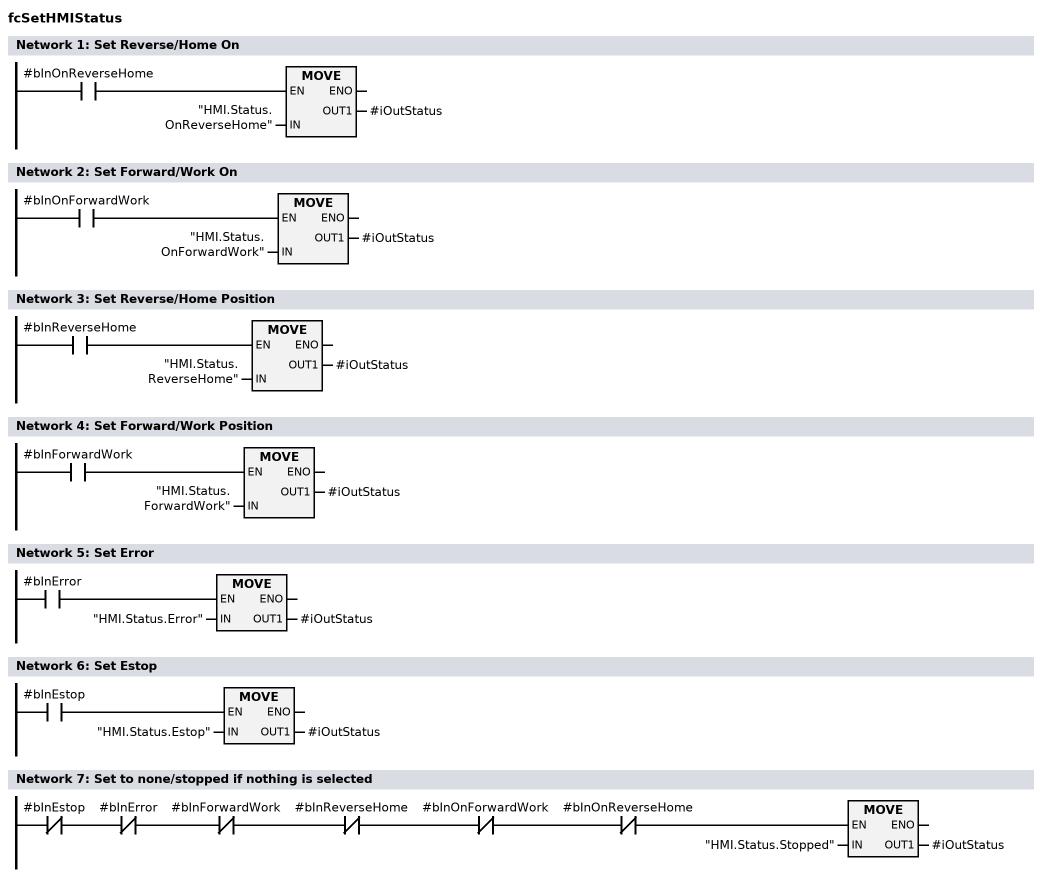
   RUNG wire#powerrail
      Contact( #bInOnReverseHome )
      Move(in := "HMI.Status.OnReverseHome", out1 => #iOutStatus)
   END_RUNG
   // the same network as SCL:
   IF #bInOnReverseHome THEN #iOutStatus := "HMI.Status.OnReverseHome"; END_IF;
END_REGION

REGION Network 2: Set Forward/Work On
   RUNG wire#powerrail
      Contact( #bInOnForwardWork )
      Move(in := "HMI.Status.OnForwardWork", out1 => #iOutStatus)
   END_RUNG
   // the same network as SCL:
   IF #bInOnForwardWork THEN #iOutStatus := "HMI.Status.OnForwardWork"; END_IF;
END_REGION

REGION Network 3: Set Reverse/Home Position
   RUNG wire#powerrail
      Contact( #bInReverseHome )
      Move(in := "HMI.Status.ReverseHome", out1 => #iOutStatus)
   END_RUNG
   // the same network as SCL:
   IF #bInReverseHome THEN #iOutStatus := "HMI.Status.ReverseHome"; END_IF;
END_REGION

REGION Network 4: Set Forward/Work Position
   RUNG wire#powerrail
      Contact( #bInForwardWork )
      Move(in := "HMI.Status.ForwardWork", out1 => #iOutStatus)
   END_RUNG
   // the same network as SCL:
   IF #bInForwardWork THEN #iOutStatus := "HMI.Status.ForwardWork"; END_IF;
END_REGION

REGION Network 5: Set Error
   RUNG wire#powerrail
      Contact( #bInError )
      Move(in := "HMI.Status.Error", out1 => #iOutStatus)
   END_RUNG
   // the same network as SCL:
   IF #bInError THEN #iOutStatus := "HMI.Status.Error"; END_IF;
END_REGION

REGION Network 6: Set Estop
   RUNG wire#powerrail
      Contact( #bInEstop )
      Move(in := "HMI.Status.Estop", out1 => #iOutStatus)
   END_RUNG
   // the same network as SCL:
   IF #bInEstop THEN #iOutStatus := "HMI.Status.Estop"; END_IF;
END_REGION

REGION Network 7: Set to none/stopped if nothing is selected
   RUNG wire#powerrail
      I_Contact( #bInEstop )
      I_Contact( #bInError )
      I_Contact( #bInForwardWork )
      I_Contact( #bInReverseHome )
      I_Contact( #bInOnForwardWork )
      I_Contact( #bInOnReverseHome )
      Move(in := "HMI.Status.Stopped", out1 => #iOutStatus)
   END_RUNG
   // the same network as SCL:
   IF NOT #bInEstop AND NOT #bInError AND NOT #bInForwardWork AND NOT #bInReverseHome AND NOT #bInOnForwardWork AND NOT #bInOnReverseHome THEN
       #iOutStatus := "HMI.Status.Stopped";
   END_IF;
END_REGION
END_FUNCTION

FUNCTION "fcSetHMIStatusGeneric" : Void   // FC1121, LAD
TITLE = Sets HMI Status
{ S7_Optimized_Access := 'FALSE' }
VERSION : 0.1
// Wrapper function for setting the HMI status of a device. 
// 
// It will display in order of priority, based on input, where Status1 > Status 2 > Status 3 > Status 4 > Status 5 > Status 6.
BEGIN

REGION Network 1: Set Status 6
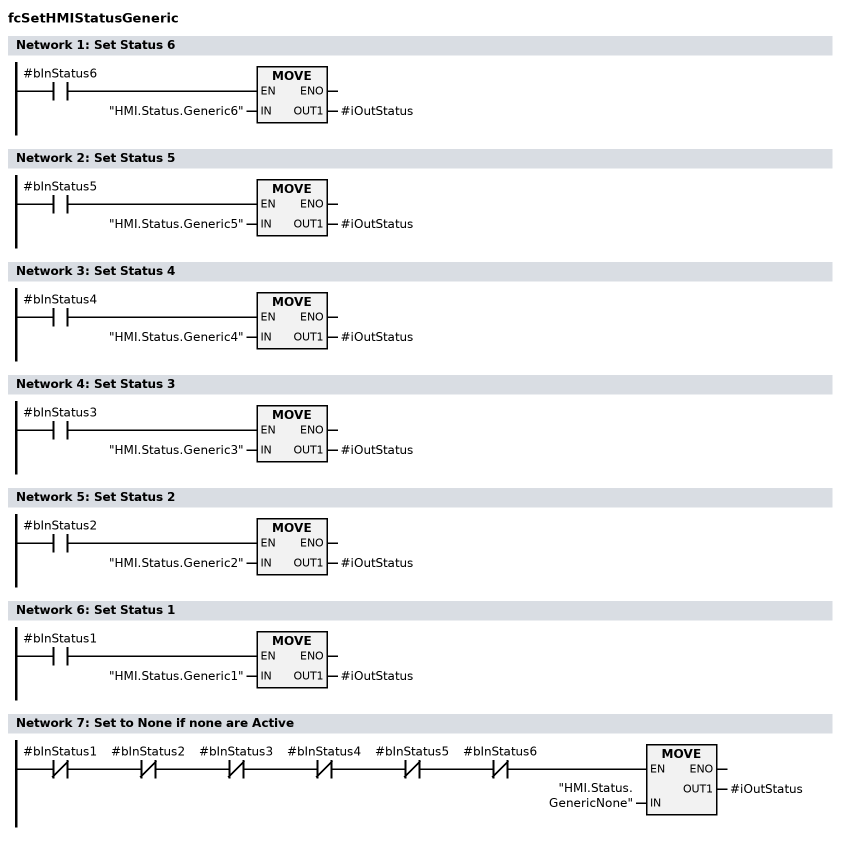
   RUNG wire#powerrail
      Contact( #bInStatus6 )
      { S7_GenerateENO := "TRUE" } Move(in := "HMI.Status.Generic6", out1 => #iOutStatus)
   END_RUNG
   // the same network as SCL:
   IF #bInStatus6 THEN #iOutStatus := "HMI.Status.Generic6"; END_IF;
END_REGION

REGION Network 2: Set Status 5
   RUNG wire#powerrail
      Contact( #bInStatus5 )
      { S7_GenerateENO := "TRUE" } Move(in := "HMI.Status.Generic5", out1 => #iOutStatus)
   END_RUNG
   // the same network as SCL:
   IF #bInStatus5 THEN #iOutStatus := "HMI.Status.Generic5"; END_IF;
END_REGION

REGION Network 3: Set Status 4
   RUNG wire#powerrail
      Contact( #bInStatus4 )
      { S7_GenerateENO := "TRUE" } Move(in := "HMI.Status.Generic4", out1 => #iOutStatus)
   END_RUNG
   // the same network as SCL:
   IF #bInStatus4 THEN #iOutStatus := "HMI.Status.Generic4"; END_IF;
END_REGION

REGION Network 4: Set Status 3
   RUNG wire#powerrail
      Contact( #bInStatus3 )
      { S7_GenerateENO := "TRUE" } Move(in := "HMI.Status.Generic3", out1 => #iOutStatus)
   END_RUNG
   // the same network as SCL:
   IF #bInStatus3 THEN #iOutStatus := "HMI.Status.Generic3"; END_IF;
END_REGION

REGION Network 5: Set Status 2
   RUNG wire#powerrail
      Contact( #bInStatus2 )
      { S7_GenerateENO := "TRUE" } Move(in := "HMI.Status.Generic2", out1 => #iOutStatus)
   END_RUNG
   // the same network as SCL:
   IF #bInStatus2 THEN #iOutStatus := "HMI.Status.Generic2"; END_IF;
END_REGION

REGION Network 6: Set Status 1
   RUNG wire#powerrail
      Contact( #bInStatus1 )
      { S7_GenerateENO := "TRUE" } Move(in := "HMI.Status.Generic1", out1 => #iOutStatus)
   END_RUNG
   // the same network as SCL:
   IF #bInStatus1 THEN #iOutStatus := "HMI.Status.Generic1"; END_IF;
END_REGION

REGION Network 7: Set to None if none are Active
   RUNG wire#powerrail
      I_Contact( #bInStatus1 )
      I_Contact( #bInStatus2 )
      I_Contact( #bInStatus3 )
      I_Contact( #bInStatus4 )
      I_Contact( #bInStatus5 )
      I_Contact( #bInStatus6 )
      { S7_GenerateENO := "TRUE" } Move(in := "HMI.Status.GenericNone", out1 => #iOutStatus)
   END_RUNG
   // the same network as SCL:
   IF NOT #bInStatus1 AND NOT #bInStatus2 AND NOT #bInStatus3 AND NOT #bInStatus4 AND NOT #bInStatus5 AND NOT #bInStatus6 THEN
       #iOutStatus := "HMI.Status.GenericNone";
   END_IF;
END_REGION
END_FUNCTION

// folder: Library Blocks/Resources/IO

FUNCTION "fcReadInput" : Void   // FC301, LAD
TITLE = Read/Scale input word
{ S7_Optimized_Access := 'FALSE' }
AUTHOR : DMC
FAMILY : IO
VERSION : 0.1
   VAR_TEMP   // added for the SCL form of the ladder/FBD networks
      _w1 : Bool;
      _w2 : Bool;
   END_VAR
BEGIN

REGION Network 1: Swap input value bytes if needed
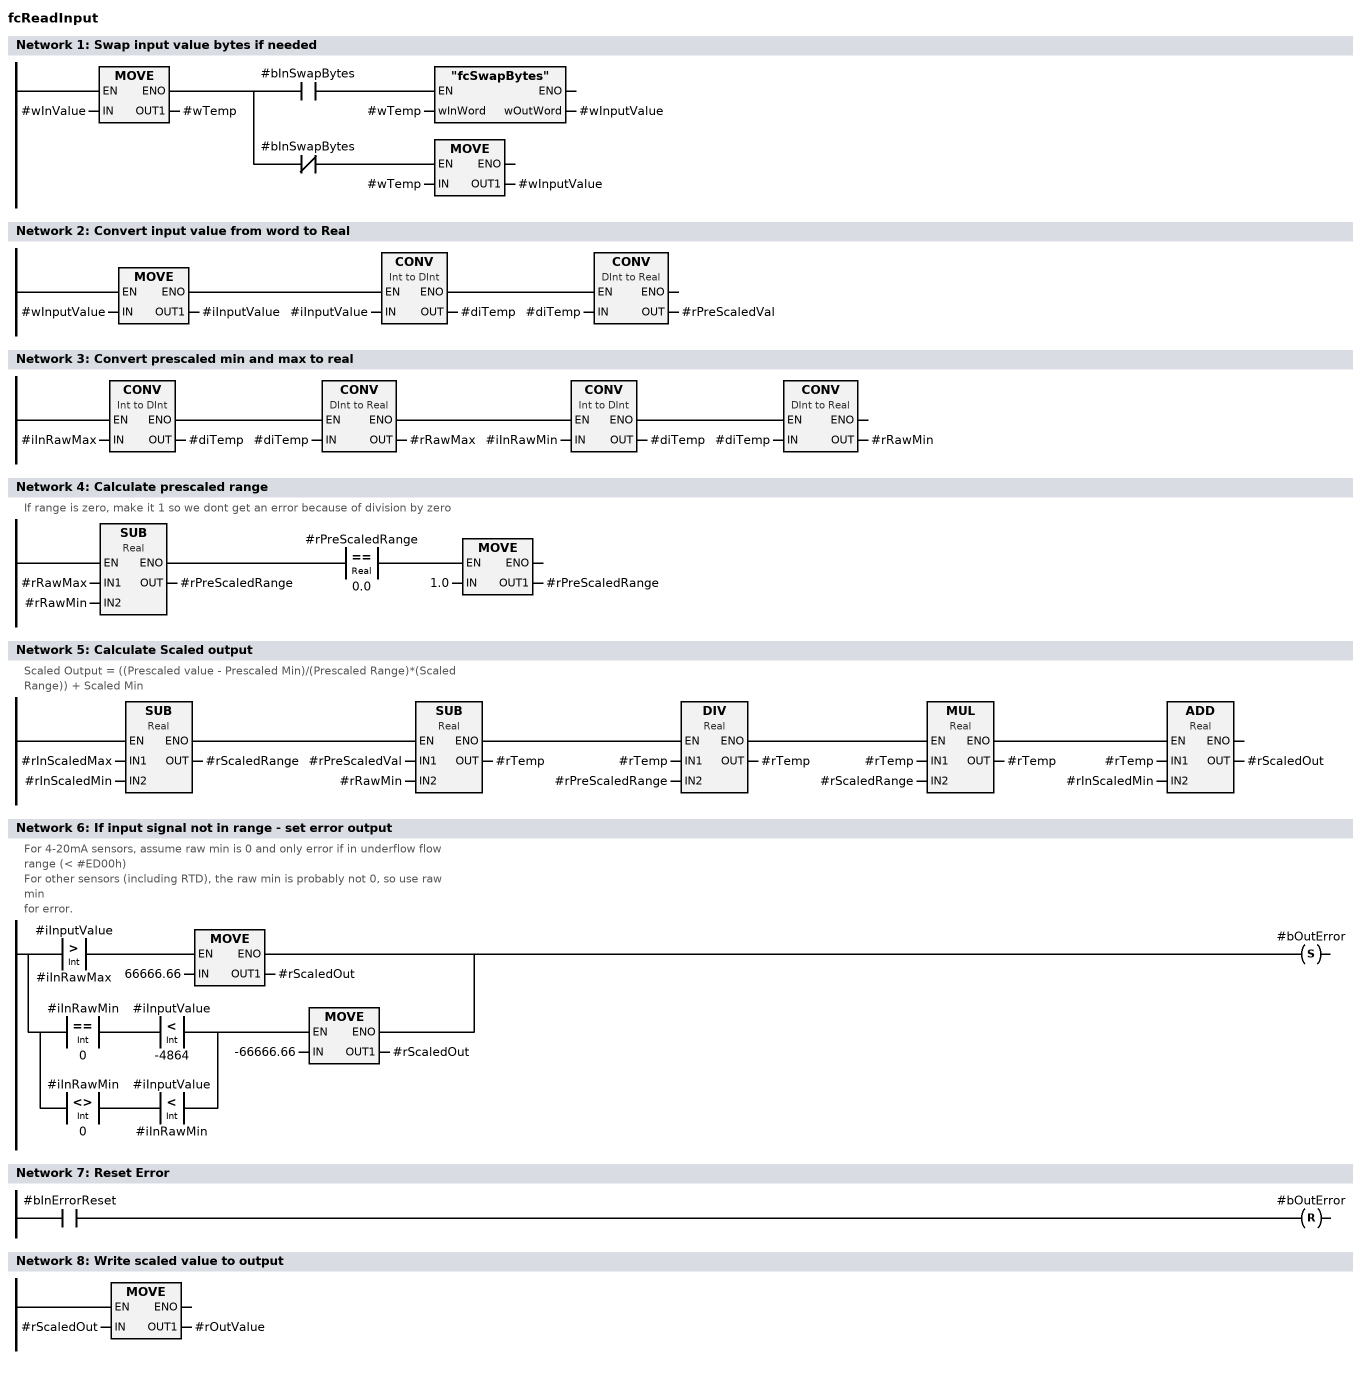
   RUNG wire#powerrail
      { S7_GenerateENO := "TRUE" } Move(in := #wInValue, out1 => #wTemp)
      wire#w1
      Contact( #bInSwapBytes )
      "fcSwapBytes"(wInWord := #wTemp, wOutWord => #wInputValue)
   END_RUNG
   RUNG wire#w1
      I_Contact( #bInSwapBytes )
      { S7_GenerateENO := "TRUE" } Move(in := #wTemp, out1 => #wInputValue)
   END_RUNG
   // the same network as SCL:
   // ENO of a box is taken as its EN; it also drops when the box reports an error
   #wTemp := #wInValue;
   IF #bInSwapBytes THEN "fcSwapBytes"(wInWord := #wTemp, wOutWord => #wInputValue); END_IF;
   IF NOT #bInSwapBytes THEN #wInputValue := #wTemp; END_IF;
END_REGION

REGION Network 2: Convert input value from word to Real
   RUNG wire#powerrail
      { S7_GenerateENO := "TRUE" } Move(in := #wInputValue, out1 => #iInputValue)
      { S7_Templates := "[SrcType := Int, DestType := DInt]"; S7_GenerateENO := "TRUE" } Convert(in := #iInputValue, out => #diTemp)
      { S7_Templates := "[SrcType := DInt, DestType := Real]"; S7_GenerateENO := "TRUE" } Convert(in := #diTemp, out => #rPreScaledVal)
   END_RUNG
   // the same network as SCL:
   // ENO of a box is taken as its EN; it also drops when the box reports an error
   #iInputValue := #wInputValue;
   #diTemp := INT_TO_DINT(#iInputValue);
   #rPreScaledVal := DINT_TO_REAL(#diTemp);
END_REGION

REGION Network 3: Convert prescaled min and max to real
   RUNG wire#powerrail
      { S7_Templates := "[SrcType := Int, DestType := DInt]"; S7_GenerateENO := "TRUE" } Convert(in := #iInRawMax, out => #diTemp)
      { S7_Templates := "[SrcType := DInt, DestType := Real]"; S7_GenerateENO := "TRUE" } Convert(in := #diTemp, out => #rRawMax)
      { S7_Templates := "[SrcType := Int, DestType := DInt]"; S7_GenerateENO := "TRUE" } Convert(in := #iInRawMin, out => #diTemp)
      { S7_Templates := "[SrcType := DInt, DestType := Real]"; S7_GenerateENO := "TRUE" } Convert(in := #diTemp, out => #rRawMin)
   END_RUNG
   // the same network as SCL:
   // ENO of a box is taken as its EN; it also drops when the box reports an error
   #diTemp := INT_TO_DINT(#iInRawMax);
   #rRawMax := DINT_TO_REAL(#diTemp);
   #diTemp := INT_TO_DINT(#iInRawMin);
   #rRawMin := DINT_TO_REAL(#diTemp);
END_REGION

REGION Network 4: Calculate prescaled range
   // If range is zero, make it 1 so we dont get an error because of division by zero
   RUNG wire#powerrail
      { S7_Templates := "SrcType := Real"; S7_GenerateENO := "TRUE" } Sub(in1 := #rRawMax, in2 := #rRawMin, out => #rPreScaledRange)
      { S7_Templates := "SrcType := Real" } EQ_Contact(in1 := #rPreScaledRange, in2 := 0.0)
      { S7_GenerateENO := "TRUE" } Move(in := 1.0, out1 => #rPreScaledRange)
   END_RUNG
   // the same network as SCL:
   // ENO of a box is taken as its EN; it also drops when the box reports an error
   #rPreScaledRange := #rRawMax - #rRawMin;
   IF #rPreScaledRange = 0.0 THEN #rPreScaledRange := 1.0; END_IF;
END_REGION

REGION Network 5: Calculate Scaled output
   // Scaled Output = ((Prescaled value - Prescaled Min)/(Prescaled Range)*(Scaled 
   // Range)) + Scaled Min
   RUNG wire#powerrail
      { S7_Templates := "SrcType := Real"; S7_GenerateENO := "TRUE" } Sub(in1 := #rInScaledMax, in2 := #rInScaledMin, out => #rScaledRange)
      { S7_Templates := "SrcType := Real"; S7_GenerateENO := "TRUE" } Sub(in1 := #rPreScaledVal, in2 := #rRawMin, out => #rTemp)
      { S7_Templates := "SrcType := Real"; S7_GenerateENO := "TRUE" } Div(in1 := #rTemp, in2 := #rPreScaledRange, out => #rTemp)
      { S7_Templates := "SrcType := Real"; S7_GenerateENO := "TRUE" } Mul(in1 := #rTemp, in2 := #rScaledRange, out => #rTemp)
      { S7_Templates := "SrcType := Real"; S7_GenerateENO := "TRUE" } Add(in1 := #rTemp, in2 := #rInScaledMin, out => #rScaledOut)
   END_RUNG
   // the same network as SCL:
   // ENO of a box is taken as its EN; it also drops when the box reports an error
   #rScaledRange := #rInScaledMax - #rInScaledMin;
   #rTemp := #rPreScaledVal - #rRawMin;
   #rTemp := #rTemp / #rPreScaledRange;
   #rTemp := #rTemp * #rScaledRange;
   #rScaledOut := #rTemp + #rInScaledMin;
END_REGION

REGION Network 6: If input signal not in range - set error output
   // For 4-20mA sensors, assume raw min is 0 and only error if in underflow flow 
   // range (< #ED00h)
   // 
   // For other sensors (including RTD), the raw min is probably not 0, so use raw 
   // min 
   // for error.
   RUNG wire#powerrail
      { S7_Templates := "SrcType := Int" } GT_Contact(in1 := #iInputValue, in2 := #iInRawMax)
      { S7_GenerateENO := "TRUE" } Move(in := 66666.66, out1 => #rScaledOut)
      wire#w1
      S_Coil( #bOutError )
   END_RUNG
   RUNG wire#powerrail
      { S7_Templates := "SrcType := Int" } EQ_Contact(in1 := #iInRawMin, in2 := 0)
      { S7_Templates := "SrcType := Int" } LT_Contact(in1 := #iInputValue, in2 := -4864)
      wire#w2
      { S7_GenerateENO := "TRUE" } Move(in := -66666.66, out1 => #rScaledOut)
   END_RUNG wire#w1
   RUNG wire#powerrail
      { S7_Templates := "SrcType := Int" } NE_Contact(in1 := #iInRawMin, in2 := 0)
      { S7_Templates := "SrcType := Int" } LT_Contact(in1 := #iInputValue, in2 := #iInRawMin)
   END_RUNG wire#w2
   // the same network as SCL:
   // ENO of a box is taken as its EN; it also drops when the box reports an error
   #_w1 := #iInputValue > #iInRawMax;
   IF #_w1 THEN #rScaledOut := 66666.66; END_IF;
   #_w2 := ((#iInRawMin = 0) AND (#iInputValue < (-4864))) OR ((#iInRawMin <> 0) AND (#iInputValue < #iInRawMin));
   IF #_w2 THEN #rScaledOut := -66666.66; END_IF;
   IF #_w1 OR #_w2 THEN #bOutError := TRUE; END_IF;
END_REGION

REGION Network 7: Reset Error
   RUNG wire#powerrail
      Contact( #bInErrorReset )
      R_Coil( #bOutError )
   END_RUNG
   // the same network as SCL:
   IF #bInErrorReset THEN #bOutError := FALSE; END_IF;
END_REGION

REGION Network 8: Write scaled value to output
   RUNG wire#powerrail
      { S7_GenerateENO := "TRUE" } Move(in := #rScaledOut, out1 => #rOutValue)
   END_RUNG
   // the same network as SCL:
   #rOutValue := #rScaledOut;
END_REGION
END_FUNCTION

FUNCTION "fcWriteOutput" : Void   // FC302, LAD
TITLE = Writes a scaled output
{ S7_Optimized_Access := 'FALSE' }
AUTHOR : DMC
FAMILY : IO
VERSION : 0.1
BEGIN

REGION Network 1: Convert raw min and max to real
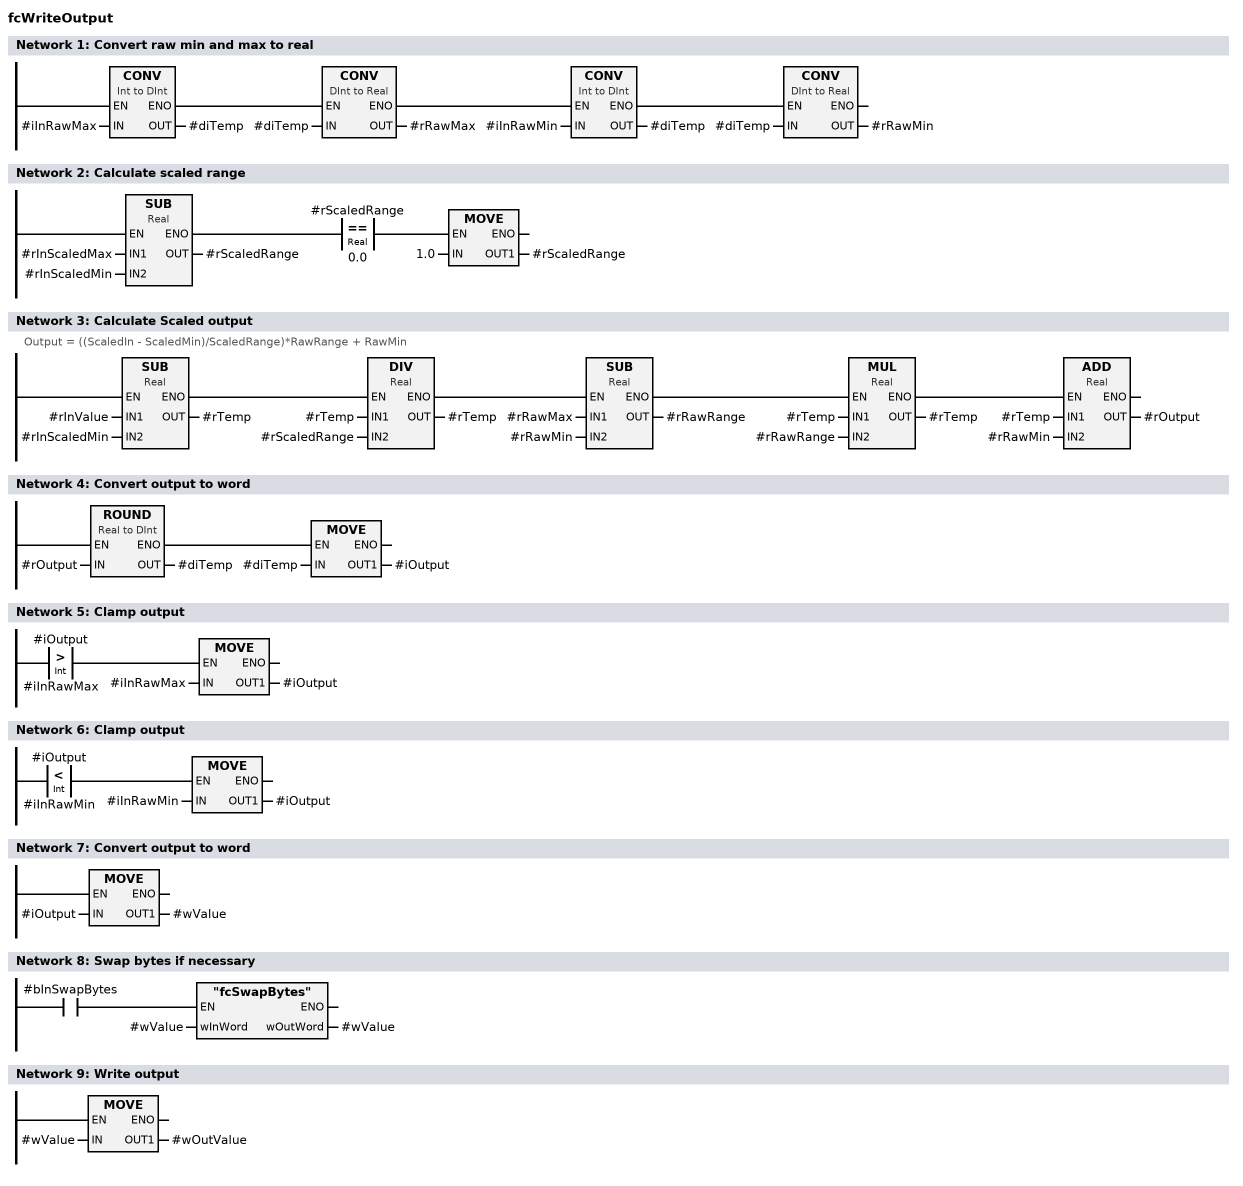
   RUNG wire#powerrail
      { S7_Templates := "[SrcType := Int, DestType := DInt]"; S7_GenerateENO := "TRUE" } Convert(in := #iInRawMax, out => #diTemp)
      { S7_Templates := "[SrcType := DInt, DestType := Real]"; S7_GenerateENO := "TRUE" } Convert(in := #diTemp, out => #rRawMax)
      { S7_Templates := "[SrcType := Int, DestType := DInt]"; S7_GenerateENO := "TRUE" } Convert(in := #iInRawMin, out => #diTemp)
      { S7_Templates := "[SrcType := DInt, DestType := Real]"; S7_GenerateENO := "TRUE" } Convert(in := #diTemp, out => #rRawMin)
   END_RUNG
   // the same network as SCL:
   // ENO of a box is taken as its EN; it also drops when the box reports an error
   #diTemp := INT_TO_DINT(#iInRawMax);
   #rRawMax := DINT_TO_REAL(#diTemp);
   #diTemp := INT_TO_DINT(#iInRawMin);
   #rRawMin := DINT_TO_REAL(#diTemp);
END_REGION

REGION Network 2: Calculate scaled range
   RUNG wire#powerrail
      { S7_Templates := "SrcType := Real"; S7_GenerateENO := "TRUE" } Sub(in1 := #rInScaledMax, in2 := #rInScaledMin, out => #rScaledRange)
      { S7_Templates := "SrcType := Real" } EQ_Contact(in1 := #rScaledRange, in2 := 0.0)
      { S7_GenerateENO := "TRUE" } Move(in := 1.0, out1 => #rScaledRange)
   END_RUNG
   // the same network as SCL:
   // ENO of a box is taken as its EN; it also drops when the box reports an error
   #rScaledRange := #rInScaledMax - #rInScaledMin;
   IF #rScaledRange = 0.0 THEN #rScaledRange := 1.0; END_IF;
END_REGION

REGION Network 3: Calculate Scaled output
   // Output = ((ScaledIn - ScaledMin)/ScaledRange)*RawRange + RawMin
   RUNG wire#powerrail
      { S7_Templates := "SrcType := Real"; S7_GenerateENO := "TRUE" } Sub(in1 := #rInValue, in2 := #rInScaledMin, out => #rTemp)
      { S7_Templates := "SrcType := Real"; S7_GenerateENO := "TRUE" } Div(in1 := #rTemp, in2 := #rScaledRange, out => #rTemp)
      { S7_Templates := "SrcType := Real"; S7_GenerateENO := "TRUE" } Sub(in1 := #rRawMax, in2 := #rRawMin, out => #rRawRange)
      { S7_Templates := "SrcType := Real"; S7_GenerateENO := "TRUE" } Mul(in1 := #rTemp, in2 := #rRawRange, out => #rTemp)
      { S7_Templates := "SrcType := Real"; S7_GenerateENO := "TRUE" } Add(in1 := #rTemp, in2 := #rRawMin, out => #rOutput)
   END_RUNG
   // the same network as SCL:
   // ENO of a box is taken as its EN; it also drops when the box reports an error
   #rTemp := #rInValue - #rInScaledMin;
   #rTemp := #rTemp / #rScaledRange;
   #rRawRange := #rRawMax - #rRawMin;
   #rTemp := #rTemp * #rRawRange;
   #rOutput := #rTemp + #rRawMin;
END_REGION

REGION Network 4: Convert output to word
   RUNG wire#powerrail
      { S7_Templates := "[SrcType := Real, DestType := DInt]"; S7_GenerateENO := "TRUE" } Round(in := #rOutput, out => #diTemp)
      { S7_GenerateENO := "TRUE" } Move(in := #diTemp, out1 => #iOutput)
   END_RUNG
   // the same network as SCL:
   // ENO of a box is taken as its EN; it also drops when the box reports an error
   #diTemp := ROUND(#rOutput);
   #iOutput := #diTemp;
END_REGION

REGION Network 5: Clamp output
   RUNG wire#powerrail
      { S7_Templates := "SrcType := Int" } GT_Contact(in1 := #iOutput, in2 := #iInRawMax)
      { S7_GenerateENO := "TRUE" } Move(in := #iInRawMax, out1 => #iOutput)
   END_RUNG
   // the same network as SCL:
   IF #iOutput > #iInRawMax THEN #iOutput := #iInRawMax; END_IF;
END_REGION

REGION Network 6: Clamp output
   RUNG wire#powerrail
      { S7_Templates := "SrcType := Int" } LT_Contact(in1 := #iOutput, in2 := #iInRawMin)
      { S7_GenerateENO := "TRUE" } Move(in := #iInRawMin, out1 => #iOutput)
   END_RUNG
   // the same network as SCL:
   IF #iOutput < #iInRawMin THEN #iOutput := #iInRawMin; END_IF;
END_REGION

REGION Network 7: Convert output to word
   RUNG wire#powerrail
      { S7_GenerateENO := "TRUE" } Move(in := #iOutput, out1 => #wValue)
   END_RUNG
   // the same network as SCL:
   #wValue := #iOutput;
END_REGION

REGION Network 8: Swap bytes if necessary
   RUNG wire#powerrail
      Contact( #bInSwapBytes )
      "fcSwapBytes"(wInWord := #wValue, wOutWord => #wValue)
   END_RUNG
   // the same network as SCL:
   IF #bInSwapBytes THEN "fcSwapBytes"(wInWord := #wValue, wOutWord => #wValue); END_IF;
END_REGION

REGION Network 9: Write output
   RUNG wire#powerrail
      { S7_GenerateENO := "TRUE" } Move(in := #wValue, out1 => #wOutValue)
   END_RUNG
   // the same network as SCL:
   #wOutValue := #wValue;
END_REGION
END_FUNCTION

FUNCTION "fcReadPIW" : Void   // FC1035, SCL
TITLE = fcReadPIW
{ S7_Optimized_Access := 'FALSE' }
AUTHOR : DMC
FAMILY : IO
NAME : RD_PIW
VERSION : 1.0
// This block read a peripheral input word
//  To use this block, feed in the address of the PIW you would like to read
//  for example: to read PIW123 you would input the number 123 to the input iPIW_Address
//  the entire word is read and output as wPIW_Value
//  Block Parameters
BEGIN


   //this reads the word from the specified peripheral input
   #wOutValue := PEEK(area := #cbyPeripheralInputArea, byteOffset := #iInAddress, dbNumber := 0);

   ENO:=TRUE;
END_FUNCTION

FUNCTION "fcWritePQW" : Void   // FC1036, SCL
TITLE = fcWritePQW
{ S7_Optimized_Access := 'FALSE' }
AUTHOR : DMC
FAMILY : IO
NAME : WR_PQW
VERSION : 1.0
// This block writes a peripheral output word
//  to use this block, enter the address of the Peripheral word and the word value.
//  for example, to set the value of PQW123 to 500, you would set iPQW_Address=123, and wPQW_Value=500
//  Block Parameters
BEGIN


   //this writes the word from the specified peripheral input
   POKE(area := #cbyPeripheralOutputArea, byteOffset := #iInAddress, dbNumber := 0, value := #wInValue);

   ENO:=TRUE;
END_FUNCTION

// folder: OBs

ORGANIZATION_BLOCK "Main"   // OB1, LAD, ProgramCycle
TITLE = "Main Program Sweep (Cycle)"
{ S7_Optimized_Access := 'FALSE' }
VERSION : 0.1
BEGIN

REGION Network 1: Master
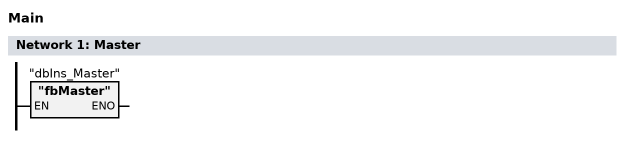
   RUNG wire#powerrail
      "dbIns_Master"()
   END_RUNG
   // the same network as SCL:
   "dbIns_Master"();   // "fbMaster"
END_REGION
END_ORGANIZATION_BLOCK

ORGANIZATION_BLOCK "Cyclic interrupt"   // OB30, LAD, CyclicInterrupt
TITLE = Cyclic Interrupt OB - 100ms
{ S7_Optimized_Access := 'FALSE' }
VERSION : 0.1
BEGIN

REGION Network 1: Call Cyclic Interrupt Function Block
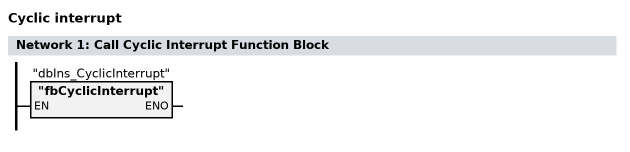
   RUNG wire#powerrail
      "dbIns_CyclicInterrupt"()
   END_RUNG
   // the same network as SCL:
   "dbIns_CyclicInterrupt"();   // "fbCyclicInterrupt"
END_REGION
END_ORGANIZATION_BLOCK

// folder: Systems/Logic

FUNCTION_BLOCK "fbWaterSystem"   // FB510, LAD
TITLE = Water System Control
{ S7_Optimized_Access := 'FALSE' }
VERSION : 0.1
   VAR_TEMP   // added for the SCL form of the ladder/FBD networks
      _w1 : Bool;
   END_VAR
BEGIN

REGION Network 1: --------------------------------------------------------- Inputs ------------------------------------------------------------------
END_REGION

REGION Network 2: Read Main Water Pump Pressure
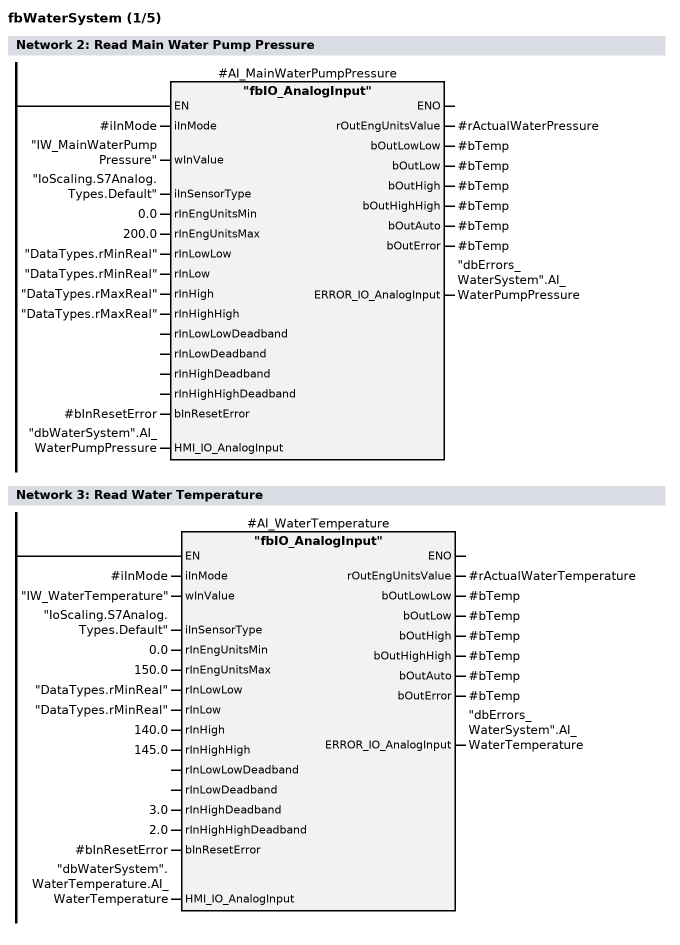
   RUNG wire#powerrail
      #AI_MainWaterPumpPressure(iInMode := #iInMode, wInValue := "IW_MainWaterPumpPressure", iInSensorType := "IoScaling.S7Analog.Types.Default", rInEngUnitsMin := 0.0, rInEngUnitsMax := 200.0, rInLowLow := "DataTypes.rMinReal", rInLow := "DataTypes.rMinReal", rInHigh := "DataTypes.rMaxReal", rInHighHigh := "DataTypes.rMaxReal", rInLowLowDeadband :=, rInLowDeadband :=, rInHighDeadband :=, rInHighHighDeadband :=, bInResetError := #bInResetError, HMI_IO_AnalogInput := "dbWaterSystem".AI_WaterPumpPressure, rOutEngUnitsValue => #rActualWaterPressure, bOutLowLow => #bTemp, bOutLow => #bTemp, bOutHigh => #bTemp, bOutHighHigh => #bTemp, bOutAuto => #bTemp, bOutError => #bTemp, ERROR_IO_AnalogInput => "dbErrors_WaterSystem".AI_WaterPumpPressure)
   END_RUNG
   // the same network as SCL:
   #AI_MainWaterPumpPressure(iInMode := #iInMode,   // "fbIO_AnalogInput"
                           wInValue := "IW_MainWaterPumpPressure",
                           iInSensorType := "IoScaling.S7Analog.Types.Default",
                           rInEngUnitsMin := 0.0,
                           rInEngUnitsMax := 200.0,
                           rInLowLow := "DataTypes.rMinReal",
                           rInLow := "DataTypes.rMinReal",
                           rInHigh := "DataTypes.rMaxReal",
                           rInHighHigh := "DataTypes.rMaxReal",
                           bInResetError := #bInResetError,
                           HMI_IO_AnalogInput := "dbWaterSystem".AI_WaterPumpPressure,
                           rOutEngUnitsValue => #rActualWaterPressure,
                           bOutLowLow => #bTemp,
                           bOutLow => #bTemp,
                           bOutHigh => #bTemp,
                           bOutHighHigh => #bTemp,
                           bOutAuto => #bTemp,
                           bOutError => #bTemp,
                           ERROR_IO_AnalogInput => "dbErrors_WaterSystem".AI_WaterPumpPressure);
END_REGION

REGION Network 3: Read Water Temperature
   RUNG wire#powerrail
      #AI_WaterTemperature(iInMode := #iInMode, wInValue := "IW_WaterTemperature", iInSensorType := "IoScaling.S7Analog.Types.Default", rInEngUnitsMin := 0.0, rInEngUnitsMax := 150.0, rInLowLow := "DataTypes.rMinReal", rInLow := "DataTypes.rMinReal", rInHigh := 140.0, rInHighHigh := 145.0, rInLowLowDeadband :=, rInLowDeadband :=, rInHighDeadband := 3.0, rInHighHighDeadband := 2.0, bInResetError := #bInResetError, HMI_IO_AnalogInput := "dbWaterSystem".WaterTemperature.AI_WaterTemperature, rOutEngUnitsValue => #rActualWaterTemperature, bOutLowLow => #bTemp, bOutLow => #bTemp, bOutHigh => #bTemp, bOutHighHigh => #bTemp, bOutAuto => #bTemp, bOutError => #bTemp, ERROR_IO_AnalogInput => "dbErrors_WaterSystem".AI_WaterTemperature)
   END_RUNG
   // the same network as SCL:
   #AI_WaterTemperature(iInMode := #iInMode,   // "fbIO_AnalogInput"
                        wInValue := "IW_WaterTemperature",
                        iInSensorType := "IoScaling.S7Analog.Types.Default",
                        rInEngUnitsMin := 0.0,
                        rInEngUnitsMax := 150.0,
                        rInLowLow := "DataTypes.rMinReal",
                        rInLow := "DataTypes.rMinReal",
                        rInHigh := 140.0,
                        rInHighHigh := 145.0,
                        rInHighDeadband := 3.0,
                        rInHighHighDeadband := 2.0,
                        bInResetError := #bInResetError,
                        HMI_IO_AnalogInput := "dbWaterSystem".WaterTemperature.AI_WaterTemperature,
                        rOutEngUnitsValue => #rActualWaterTemperature,
                        bOutLowLow => #bTemp,
                        bOutLow => #bTemp,
                        bOutHigh => #bTemp,
                        bOutHighHigh => #bTemp,
                        bOutAuto => #bTemp,
                        bOutError => #bTemp,
                        ERROR_IO_AnalogInput => "dbErrors_WaterSystem".AI_WaterTemperature);
END_REGION

REGION Network 4: --------------------------------------------------- System Logic ------------------------------------------------------------
END_REGION

REGION Network 5: Main Water Pump Interlock
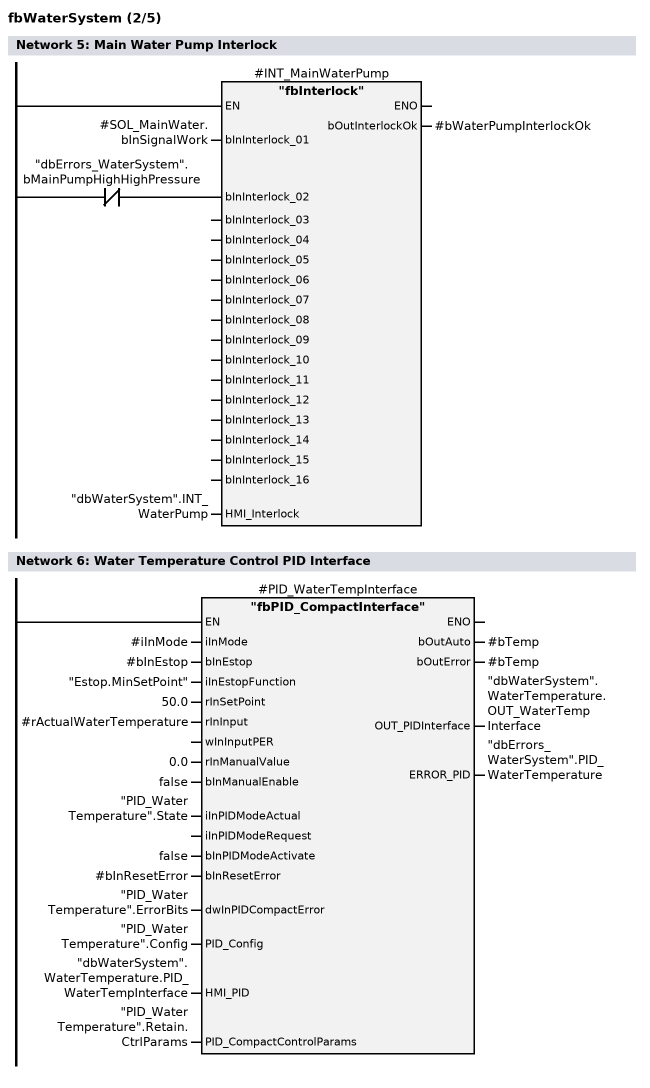
   RUNG wire#powerrail
      #INT_MainWaterPump(bInInterlock_02 := wire#w1, bInInterlock_01 := #SOL_MainWater.bInSignalWork, bInInterlock_03 :=, bInInterlock_04 :=, bInInterlock_05 :=, bInInterlock_06 :=, bInInterlock_07 :=, bInInterlock_08 :=, bInInterlock_09 :=, bInInterlock_10 :=, bInInterlock_11 :=, bInInterlock_12 :=, bInInterlock_13 :=, bInInterlock_14 :=, bInInterlock_15 :=, bInInterlock_16 :=, HMI_Interlock := "dbWaterSystem".INT_WaterPump, bOutInterlockOk => #bWaterPumpInterlockOk)
   END_RUNG
   RUNG wire#powerrail
      I_Contact( "dbErrors_WaterSystem".bMainPumpHighHighPressure )
   END_RUNG wire#w1
   // the same network as SCL:
   #INT_MainWaterPump(bInInterlock_01 := #SOL_MainWater.bInSignalWork,   // "fbInterlock"
                      bInInterlock_02 := NOT "dbErrors_WaterSystem".bMainPumpHighHighPressure,
                      HMI_Interlock := "dbWaterSystem".INT_WaterPump,
                      bOutInterlockOk => #bWaterPumpInterlockOk);
END_REGION

REGION Network 6: Water Temperature Control PID Interface
   RUNG wire#powerrail
      #PID_WaterTempInterface(iInMode := #iInMode, bInEstop := #bInEstop, iInEstopFunction := "Estop.MinSetPoint", rInSetPoint := 50.0, rInInput := #rActualWaterTemperature, wInInputPER :=, rInManualValue := 0.0, bInManualEnable := false, iInPIDModeActual := "PID_WaterTemperature".State, iInPIDModeRequest :=, bInPIDModeActivate := false, bInResetError := #bInResetError, dwInPIDCompactError := "PID_WaterTemperature".ErrorBits, PID_Config := "PID_WaterTemperature".Config, HMI_PID := "dbWaterSystem".WaterTemperature.PID_WaterTempInterface, PID_CompactControlParams := "PID_WaterTemperature".Retain.CtrlParams, bOutAuto => #bTemp, bOutError => #bTemp, OUT_PIDInterface => "dbWaterSystem".WaterTemperature.OUT_WaterTempInterface, ERROR_PID => "dbErrors_WaterSystem".PID_WaterTemperature)
   END_RUNG
   // the same network as SCL:
   #PID_WaterTempInterface(iInMode := #iInMode,   // "fbPID_CompactInterface"
                           bInEstop := #bInEstop,
                           iInEstopFunction := "Estop.MinSetPoint",
                           rInSetPoint := 50.0,
                           rInInput := #rActualWaterTemperature,
                           rInManualValue := 0.0,
                           bInManualEnable := false,
                           iInPIDModeActual := "PID_WaterTemperature".State,
                           bInPIDModeActivate := false,
                           bInResetError := #bInResetError,
                           dwInPIDCompactError := "PID_WaterTemperature".ErrorBits,
                           PID_Config := "PID_WaterTemperature".Config,
                           HMI_PID := "dbWaterSystem".WaterTemperature.PID_WaterTempInterface,
                           PID_CompactControlParams := "PID_WaterTemperature".Retain.CtrlParams,
                           bOutAuto => #bTemp,
                           bOutError => #bTemp,
                           OUT_PIDInterface => "dbWaterSystem".WaterTemperature.OUT_WaterTempInterface,
                           ERROR_PID => "dbErrors_WaterSystem".PID_WaterTemperature);
END_REGION

REGION Network 7: Determine steam valve and cooling coil set points
   // If the PID output is greater than zero, we want to open the steam valve
   // If it is less than zero, we want to increase the cooling coil
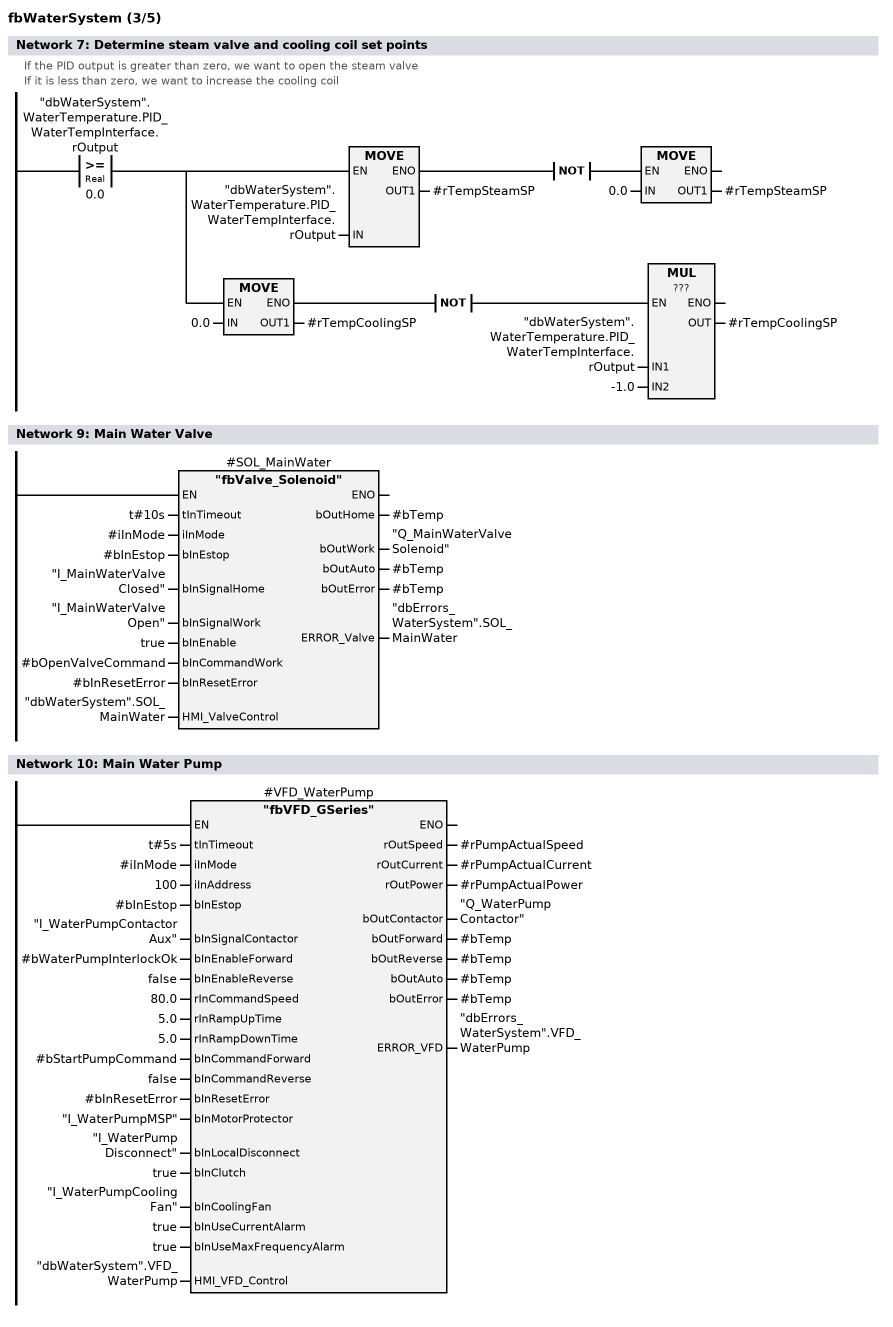
   RUNG wire#powerrail
      { S7_Templates := "SrcType := Real" } GE_Contact(in1 := "dbWaterSystem".WaterTemperature.PID_WaterTempInterface.rOutput, in2 := 0.0)
      wire#w1
      Move(in := "dbWaterSystem".WaterTemperature.PID_WaterTempInterface.rOutput, out1 => #rTempSteamSP)
      Not()
      Move(in := 0.0, out1 => #rTempSteamSP)
   END_RUNG
   RUNG wire#w1
      Move(in := 0.0, out1 => #rTempCoolingSP)
      Not()
      { S7_Templates := "SrcType := ???" } Mul(in1 := "dbWaterSystem".WaterTemperature.PID_WaterTempInterface.rOutput, in2 := -1.0, out => #rTempCoolingSP)
   END_RUNG
   // the same network as SCL:
   #_w1 := "dbWaterSystem".WaterTemperature.PID_WaterTempInterface.rOutput >= 0.0;
   IF #_w1 THEN #rTempSteamSP := "dbWaterSystem".WaterTemperature.PID_WaterTempInterface.rOutput; END_IF;
   IF NOT #_w1 THEN #rTempSteamSP := 0.0; END_IF;
   IF #_w1 THEN #rTempCoolingSP := 0.0; END_IF;
   IF NOT #_w1 THEN
       #rTempCoolingSP := "dbWaterSystem".WaterTemperature.PID_WaterTempInterface.rOutput * (-1.0);
   END_IF;
END_REGION

REGION Network 8: -------------------------------------------------------- Devices -----------------------------------------------------------------
END_REGION

REGION Network 9: Main Water Valve
   RUNG wire#powerrail
      #SOL_MainWater(tInTimeout := t#10s, iInMode := #iInMode, bInEstop := #bInEstop, bInSignalHome := "I_MainWaterValveClosed", bInSignalWork := "I_MainWaterValveOpen", bInEnable := true, bInCommandWork := #bOpenValveCommand, bInResetError := #bInResetError, HMI_ValveControl := "dbWaterSystem".SOL_MainWater, bOutHome => #bTemp, bOutWork => "Q_MainWaterValveSolenoid", bOutAuto => #bTemp, bOutError => #bTemp, ERROR_Valve => "dbErrors_WaterSystem".SOL_MainWater)
   END_RUNG
   // the same network as SCL:
   #SOL_MainWater(tInTimeout := t#10s,   // "fbValve_Solenoid"
                  iInMode := #iInMode,
                  bInEstop := #bInEstop,
                  bInSignalHome := "I_MainWaterValveClosed",
                  bInSignalWork := "I_MainWaterValveOpen",
                  bInEnable := true,
                  bInCommandWork := #bOpenValveCommand,
                  bInResetError := #bInResetError,
                  HMI_ValveControl := "dbWaterSystem".SOL_MainWater,
                  bOutHome => #bTemp,
                  bOutWork => "Q_MainWaterValveSolenoid",
                  bOutAuto => #bTemp,
                  bOutError => #bTemp,
                  ERROR_Valve => "dbErrors_WaterSystem".SOL_MainWater);
END_REGION
